REGION Network 15: Position Carrier Control First Carrier in Accumulation Zone
   RUNG wire#powerrail
      Contact( "EMS".Zone[#Zone].AccumZone )
      wire#w1
      I_Contact( "EMS".Zone[#NextZone].ZoneFull )
      wire#w2
      Move(in := #NextStopPosition, out1 => #TrafficCopCarrierZnBuffer[#ZonePos].CommandPos)
      wire#w3
      I_Contact( "EMS".Zone[#Zone].FinePosStopZone )
      Sub(in1 := #TrafficCopCarrierZnBuffer[#ZonePos].CommandPos, in2 := "EMS".CoarsePositionTolerance, out => #TrafficCopCarrierZnBuffer[#ZonePos].CommandPosLowLimit)
      Add(in1 := #TrafficCopCarrierZnBuffer[#ZonePos].CommandPos, in2 := "EMS".CoarsePositionTolerance, out => #TrafficCopCarrierZnBuffer[#ZonePos].CommandPosHighLimit)
   END_RUNG
   RUNG wire#w1
      { S7_Templates := "SrcType := DInt" } LT_Contact(in1 := "EMS".Zone[#Zone].CarrierZnStatus[#ZonePos].Position, in2 := #EndPos_LowLimit)
   END_RUNG wire#w2
   RUNG wire#w1
      { S7_Templates := "SrcType := DInt" } GE_Contact(in1 := "EMS".Zone[#Zone].CarrierZnStatus[#ZonePos].Position, in2 := #EndPos_LowLimit)
      { S7_Templates := "SrcType := DInt" } LE_Contact(in1 := "EMS".Zone[#Zone].CarrierZnStatus[#ZonePos].Position, in2 := #EndPos_HighLimit)
      { S7_Templates := "SrcType := Word" } EQ_Contact(in1 := "EMS".Zone[#NextZone].CarrierZnStatus[1].CarrierNumber, in2 := 0)
   END_RUNG wire#w2
   RUNG wire#powerrail
      Contact( "EMS".Zone[#Zone].ProductionZone )
      { S7_Templates := "SrcType := DInt" } LT_Contact(in1 := "EMS".Zone[#Zone].CarrierZnStatus[#ZonePos].Position, in2 := #ClrOfStopPos_LowLimit)
      Move(in := #ClearOfStopPos, out1 => #TrafficCopCarrierZnBuffer[#ZonePos].CommandPos)
   END_RUNG wire#w3
   RUNG wire#w3
      Contact( "EMS".Zone[#Zone].FinePosStopZone )
      Sub(in1 := #TrafficCopCarrierZnBuffer[#ZonePos].CommandPos, in2 := "EMS".FinePositionTolerance, out => #TrafficCopCarrierZnBuffer[#ZonePos].CommandPosLowLimit)
      Add(in1 := #TrafficCopCarrierZnBuffer[#ZonePos].CommandPos, in2 := "EMS".FinePositionTolerance, out => #TrafficCopCarrierZnBuffer[#ZonePos].CommandPosHighLimit)
   END_RUNG
   // the same network as SCL:
   #_w1 := "EMS".Zone[#Zone].AccumZone AND (NOT "EMS".Zone[#NextZone].ZoneFull OR ("EMS".Zone[#Zone].CarrierZnStatus[#ZonePos].Position < #EndPos_LowLimit) OR (("EMS".Zone[#Zone].CarrierZnStatus[#ZonePos].Position >= #EndPos_LowLimit) AND ("EMS".Zone[#Zone].CarrierZnStatus[#ZonePos].Position <= #EndPos_HighLimit) AND ("EMS".Zone[#NextZone].CarrierZnStatus[1].CarrierNumber = 0)));
   IF #_w1 THEN #TrafficCopCarrierZnBuffer[#ZonePos].CommandPos := #NextStopPosition; END_IF;
   #_w2 := "EMS".Zone[#Zone].ProductionZone AND ("EMS".Zone[#Zone].CarrierZnStatus[#ZonePos].Position < #ClrOfStopPos_LowLimit);
   IF #_w2 THEN #TrafficCopCarrierZnBuffer[#ZonePos].CommandPos := #ClearOfStopPos; END_IF;
   #_w3 := #_w1 OR #_w2;
   IF #_w3 AND NOT "EMS".Zone[#Zone].FinePosStopZone THEN
       #TrafficCopCarrierZnBuffer[#ZonePos].CommandPosLowLimit := #TrafficCopCarrierZnBuffer[#ZonePos].CommandPos - "EMS".CoarsePositionTolerance;
       #TrafficCopCarrierZnBuffer[#ZonePos].CommandPosHighLimit := #TrafficCopCarrierZnBuffer[#ZonePos].CommandPos + "EMS".CoarsePositionTolerance;
   END_IF;
   IF #_w3 AND "EMS".Zone[#Zone].FinePosStopZone THEN
       #TrafficCopCarrierZnBuffer[#ZonePos].CommandPosLowLimit := #TrafficCopCarrierZnBuffer[#ZonePos].CommandPos - "EMS".FinePositionTolerance;
       #TrafficCopCarrierZnBuffer[#ZonePos].CommandPosHighLimit := #TrafficCopCarrierZnBuffer[#ZonePos].CommandPos + "EMS".FinePositionTolerance;
   END_IF;
END_REGION

REGION Network 16: Position Carrier Control First Carrier in Production Zone
   // Control of First Carrier in Zone Closest to end position/Stop.  Move command is issued to carrier. Carrier will move in auto.
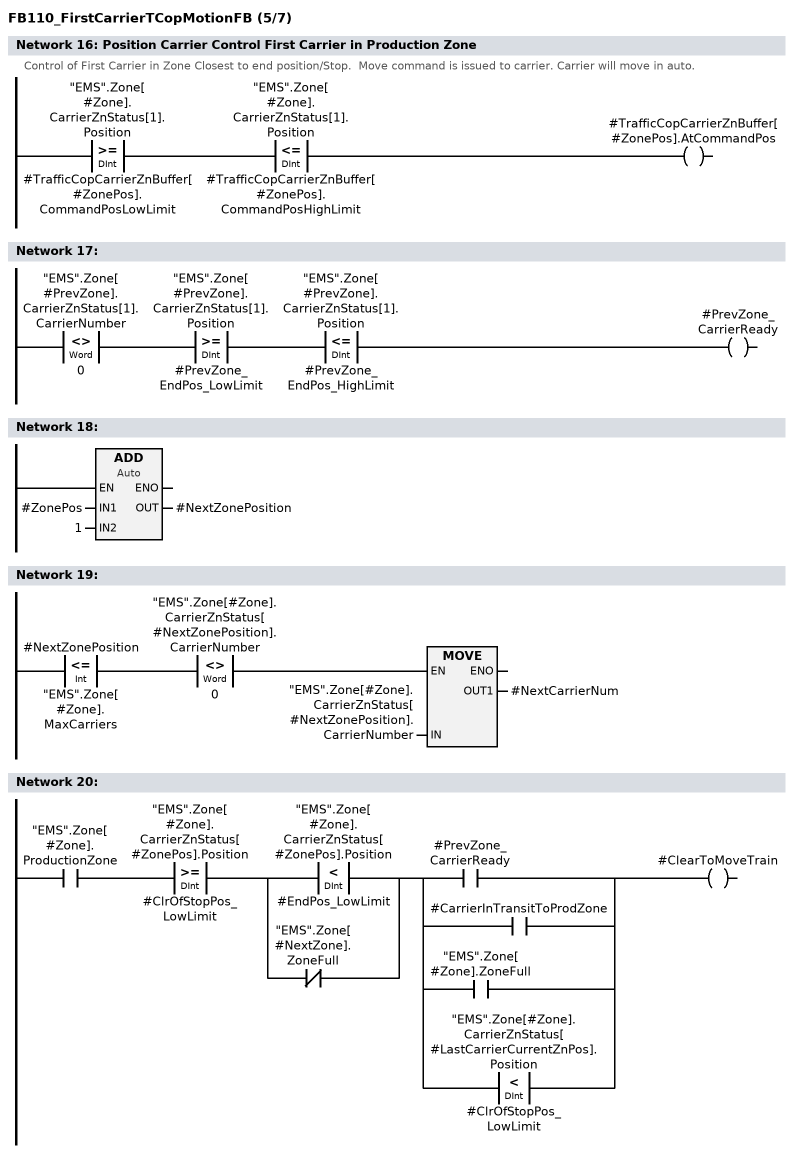
   RUNG wire#powerrail
      { S7_Templates := "SrcType := DInt" } GE_Contact(in1 := "EMS".Zone[#Zone].CarrierZnStatus[1].Position, in2 := #TrafficCopCarrierZnBuffer[#ZonePos].CommandPosLowLimit)
      { S7_Templates := "SrcType := DInt" } LE_Contact(in1 := "EMS".Zone[#Zone].CarrierZnStatus[1].Position, in2 := #TrafficCopCarrierZnBuffer[#ZonePos].CommandPosHighLimit)
      Coil( #TrafficCopCarrierZnBuffer[#ZonePos].AtCommandPos )
   END_RUNG
   // the same network as SCL:
   #TrafficCopCarrierZnBuffer[#ZonePos].AtCommandPos := ("EMS".Zone[#Zone].CarrierZnStatus[1].Position >= #TrafficCopCarrierZnBuffer[#ZonePos].CommandPosLowLimit) AND ("EMS".Zone[#Zone].CarrierZnStatus[1].Position <= #TrafficCopCarrierZnBuffer[#ZonePos].CommandPosHighLimit);
END_REGION

REGION Network 17
   RUNG wire#powerrail
      { S7_Templates := "SrcType := Word" } NE_Contact(in1 := "EMS".Zone[#PrevZone].CarrierZnStatus[1].CarrierNumber, in2 := 0)
      { S7_Templates := "SrcType := DInt" } GE_Contact(in1 := "EMS".Zone[#PrevZone].CarrierZnStatus[1].Position, in2 := #PrevZone_EndPos_LowLimit)
      { S7_Templates := "SrcType := DInt" } LE_Contact(in1 := "EMS".Zone[#PrevZone].CarrierZnStatus[1].Position, in2 := #PrevZone_EndPos_HighLimit)
      Coil( #PrevZone_CarrierReady )
   END_RUNG
   // the same network as SCL:
   #PrevZone_CarrierReady := ("EMS".Zone[#PrevZone].CarrierZnStatus[1].CarrierNumber <> 0) AND ("EMS".Zone[#PrevZone].CarrierZnStatus[1].Position >= #PrevZone_EndPos_LowLimit) AND ("EMS".Zone[#PrevZone].CarrierZnStatus[1].Position <= #PrevZone_EndPos_HighLimit);
END_REGION

REGION Network 18
   RUNG wire#powerrail
      Add(in1 := #ZonePos, in2 := 1, out => #NextZonePosition)
   END_RUNG
   // the same network as SCL:
   #NextZonePosition := #ZonePos + 1;
END_REGION

REGION Network 19
   RUNG wire#powerrail
      { S7_Templates := "SrcType := Int" } LE_Contact(in1 := #NextZonePosition, in2 := "EMS".Zone[#Zone].MaxCarriers)
      { S7_Templates := "SrcType := Word" } NE_Contact(in1 := "EMS".Zone[#Zone].CarrierZnStatus[#NextZonePosition].CarrierNumber, in2 := 0)
      Move(in := "EMS".Zone[#Zone].CarrierZnStatus[#NextZonePosition].CarrierNumber, out1 => #NextCarrierNum)
   END_RUNG
   // the same network as SCL:
   IF (#NextZonePosition <= "EMS".Zone[#Zone].MaxCarriers) AND ("EMS".Zone[#Zone].CarrierZnStatus[#NextZonePosition].CarrierNumber <> 0) THEN
       #NextCarrierNum := "EMS".Zone[#Zone].CarrierZnStatus[#NextZonePosition].CarrierNumber;
   END_IF;
END_REGION

REGION Network 20
   RUNG wire#powerrail
      Contact( "EMS".Zone[#Zone].ProductionZone )
      { S7_Templates := "SrcType := DInt" } GE_Contact(in1 := "EMS".Zone[#Zone].CarrierZnStatus[#ZonePos].Position, in2 := #ClrOfStopPos_LowLimit)
      wire#w1
      { S7_Templates := "SrcType := DInt" } LT_Contact(in1 := "EMS".Zone[#Zone].CarrierZnStatus[#ZonePos].Position, in2 := #EndPos_LowLimit)
      wire#w2
      Contact( #PrevZone_CarrierReady )
      wire#w3
      Coil( #ClearToMoveTrain )
   END_RUNG
   RUNG wire#w1
      I_Contact( "EMS".Zone[#NextZone].ZoneFull )
   END_RUNG wire#w2
   RUNG wire#w2
      Contact( #CarrierInTransitToProdZone )
   END_RUNG wire#w3
   RUNG wire#w2
      Contact( "EMS".Zone[#Zone].ZoneFull )
   END_RUNG wire#w3
   RUNG wire#w2
      { S7_Templates := "SrcType := DInt" } LT_Contact(in1 := "EMS".Zone[#Zone].CarrierZnStatus[#LastCarrierCurrentZnPos].Position, in2 := #ClrOfStopPos_LowLimit)
   END_RUNG wire#w3
   // the same network as SCL:
   #ClearToMoveTrain := "EMS".Zone[#Zone].ProductionZone AND ("EMS".Zone[#Zone].CarrierZnStatus[#ZonePos].Position >= #ClrOfStopPos_LowLimit) AND (("EMS".Zone[#Zone].CarrierZnStatus[#ZonePos].Position < #EndPos_LowLimit) OR NOT "EMS".Zone[#NextZone].ZoneFull) AND (#PrevZone_CarrierReady OR #CarrierInTransitToProdZone OR "EMS".Zone[#Zone].ZoneFull OR ("EMS".Zone[#Zone].CarrierZnStatus[#LastCarrierCurrentZnPos].Position < #ClrOfStopPos_LowLimit));
END_REGION

REGION Network 21
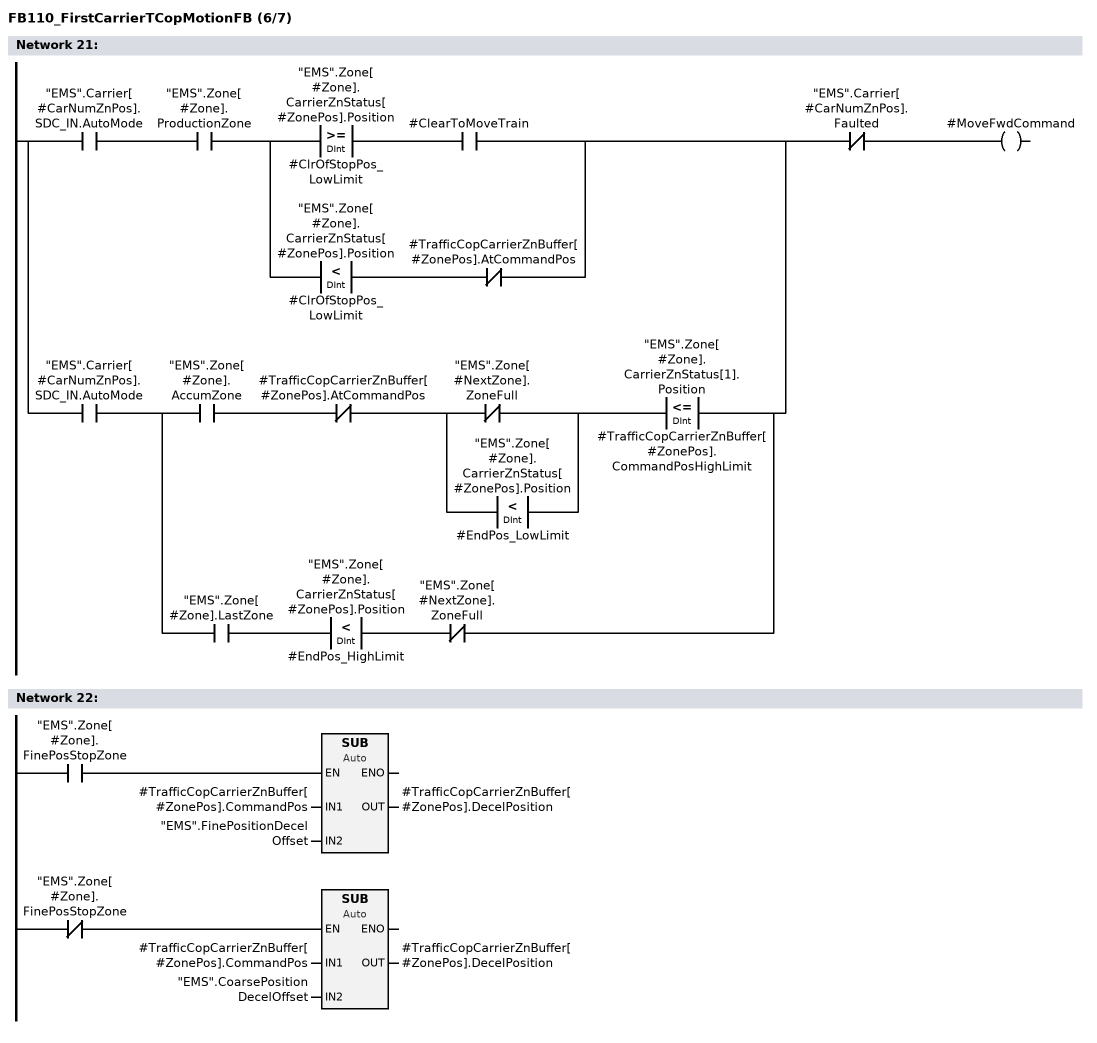
   RUNG wire#powerrail
      Contact( "EMS".Carrier[#CarNumZnPos].SDC_IN.AutoMode )
      Contact( "EMS".Zone[#Zone].ProductionZone )
      wire#w1
      { S7_Templates := "SrcType := DInt" } GE_Contact(in1 := "EMS".Zone[#Zone].CarrierZnStatus[#ZonePos].Position, in2 := #ClrOfStopPos_LowLimit)
      Contact( #ClearToMoveTrain )
      wire#w2
      I_Contact( "EMS".Carrier[#CarNumZnPos].Faulted )
      Coil( #MoveFwdCommand )
   END_RUNG
   RUNG wire#w1
      { S7_Templates := "SrcType := DInt" } LT_Contact(in1 := "EMS".Zone[#Zone].CarrierZnStatus[#ZonePos].Position, in2 := #ClrOfStopPos_LowLimit)
      I_Contact( #TrafficCopCarrierZnBuffer[#ZonePos].AtCommandPos )
   END_RUNG wire#w2
   RUNG wire#powerrail
      Contact( "EMS".Carrier[#CarNumZnPos].SDC_IN.AutoMode )
      wire#w3
      Contact( "EMS".Zone[#Zone].AccumZone )
      I_Contact( #TrafficCopCarrierZnBuffer[#ZonePos].AtCommandPos )
      wire#w4
      I_Contact( "EMS".Zone[#NextZone].ZoneFull )
      wire#w5
      { S7_Templates := "SrcType := DInt" } LE_Contact(in1 := "EMS".Zone[#Zone].CarrierZnStatus[1].Position, in2 := #TrafficCopCarrierZnBuffer[#ZonePos].CommandPosHighLimit)
   END_RUNG wire#w2
   RUNG wire#w4
      { S7_Templates := "SrcType := DInt" } LT_Contact(in1 := "EMS".Zone[#Zone].CarrierZnStatus[#ZonePos].Position, in2 := #EndPos_LowLimit)
   END_RUNG wire#w5
   RUNG wire#w3
      Contact( "EMS".Zone[#Zone].LastZone )
      { S7_Templates := "SrcType := DInt" } LT_Contact(in1 := "EMS".Zone[#Zone].CarrierZnStatus[#ZonePos].Position, in2 := #EndPos_HighLimit)
      I_Contact( "EMS".Zone[#NextZone].ZoneFull )
   END_RUNG wire#w2
   // the same network as SCL:
   #MoveFwdCommand := (("EMS".Carrier[#CarNumZnPos].SDC_IN.AutoMode AND "EMS".Zone[#Zone].ProductionZone AND ((("EMS".Zone[#Zone].CarrierZnStatus[#ZonePos].Position >= #ClrOfStopPos_LowLimit) AND #ClearToMoveTrain) OR (("EMS".Zone[#Zone].CarrierZnStatus[#ZonePos].Position < #ClrOfStopPos_LowLimit) AND NOT #TrafficCopCarrierZnBuffer[#ZonePos].AtCommandPos))) OR ("EMS".Carrier[#CarNumZnPos].SDC_IN.AutoMode AND (("EMS".Zone[#Zone].AccumZone AND NOT #TrafficCopCarrierZnBuffer[#ZonePos].AtCommandPos AND (NOT "EMS".Zone[#NextZone].ZoneFull OR ("EMS".Zone[#Zone].CarrierZnStatus[#ZonePos].Position < #EndPos_LowLimit)) AND ("EMS".Zone[#Zone].CarrierZnStatus[1].Position <= #TrafficCopCarrierZnBuffer[#ZonePos].CommandPosHighLimit)) OR ("EMS".Zone[#Zone].LastZone AND ("EMS".Zone[#Zone].CarrierZnStatus[#ZonePos].Position < #EndPos_HighLimit) AND NOT "EMS".Zone[#NextZone].ZoneFull)))) AND NOT "EMS".Carrier[#CarNumZnPos].Faulted;
END_REGION

REGION Network 22
   RUNG wire#powerrail
      Contact( "EMS".Zone[#Zone].FinePosStopZone )
      Sub(in1 := #TrafficCopCarrierZnBuffer[#ZonePos].CommandPos, in2 := "EMS".FinePositionDecelOffset, out => #TrafficCopCarrierZnBuffer[#ZonePos].DecelPosition)
   END_RUNG
   RUNG wire#powerrail
      I_Contact( "EMS".Zone[#Zone].FinePosStopZone )
      Sub(in1 := #TrafficCopCarrierZnBuffer[#ZonePos].CommandPos, in2 := "EMS".CoarsePositionDecelOffset, out => #TrafficCopCarrierZnBuffer[#ZonePos].DecelPosition)
   END_RUNG
   // the same network as SCL:
   IF "EMS".Zone[#Zone].FinePosStopZone THEN
       #TrafficCopCarrierZnBuffer[#ZonePos].DecelPosition := #TrafficCopCarrierZnBuffer[#ZonePos].CommandPos - "EMS".FinePositionDecelOffset;
   END_IF;
   IF NOT "EMS".Zone[#Zone].FinePosStopZone THEN
       #TrafficCopCarrierZnBuffer[#ZonePos].DecelPosition := #TrafficCopCarrierZnBuffer[#ZonePos].CommandPos - "EMS".CoarsePositionDecelOffset;
   END_IF;
END_REGION

REGION Network 23
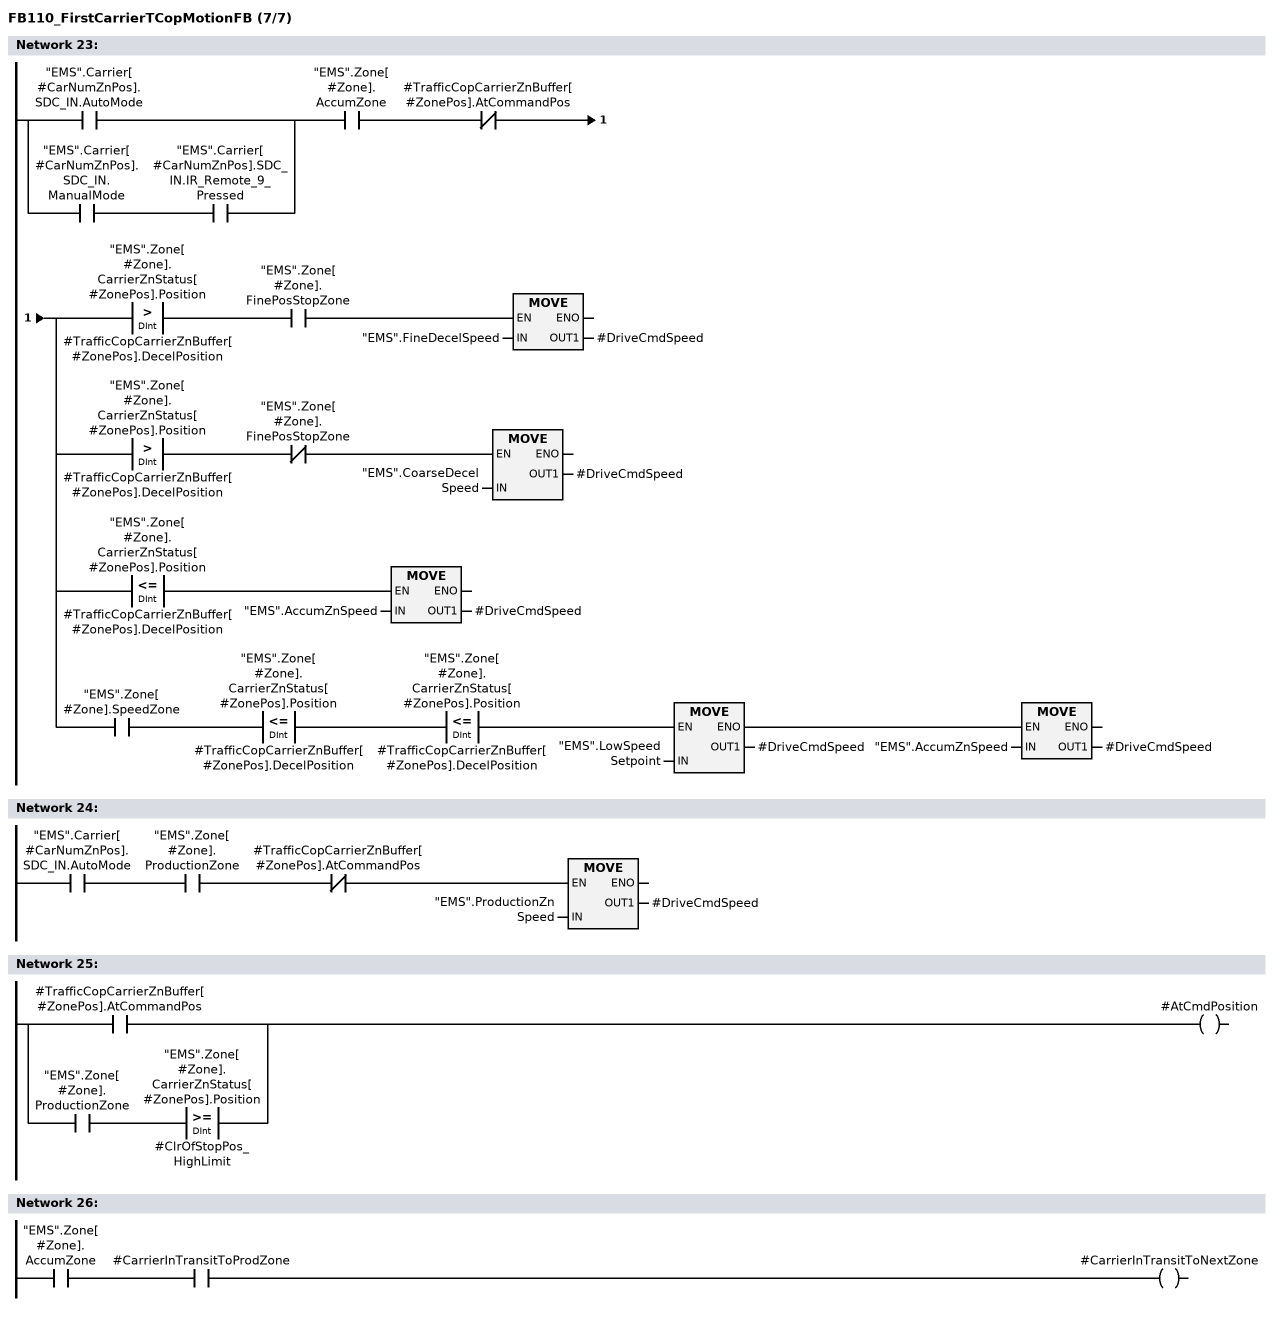
   RUNG wire#powerrail
      Contact( "EMS".Carrier[#CarNumZnPos].SDC_IN.AutoMode )
      wire#w1
      Contact( "EMS".Zone[#Zone].AccumZone )
      I_Contact( #TrafficCopCarrierZnBuffer[#ZonePos].AtCommandPos )
      wire#w2
      { S7_Templates := "SrcType := DInt" } GT_Contact(in1 := "EMS".Zone[#Zone].CarrierZnStatus[#ZonePos].Position, in2 := #TrafficCopCarrierZnBuffer[#ZonePos].DecelPosition)
      Contact( "EMS".Zone[#Zone].FinePosStopZone )
      Move(in := "EMS".FineDecelSpeed, out1 => #DriveCmdSpeed)
   END_RUNG
   RUNG wire#powerrail
      Contact( "EMS".Carrier[#CarNumZnPos].SDC_IN.ManualMode )
      Contact( "EMS".Carrier[#CarNumZnPos].SDC_IN.IR_Remote_9_Pressed )
   END_RUNG wire#w1
   RUNG wire#w2
      { S7_Templates := "SrcType := DInt" } GT_Contact(in1 := "EMS".Zone[#Zone].CarrierZnStatus[#ZonePos].Position, in2 := #TrafficCopCarrierZnBuffer[#ZonePos].DecelPosition)
      I_Contact( "EMS".Zone[#Zone].FinePosStopZone )
      Move(in := "EMS".CoarseDecelSpeed, out1 => #DriveCmdSpeed)
   END_RUNG
   RUNG wire#w2
      { S7_Templates := "SrcType := DInt" } LE_Contact(in1 := "EMS".Zone[#Zone].CarrierZnStatus[#ZonePos].Position, in2 := #TrafficCopCarrierZnBuffer[#ZonePos].DecelPosition)
      Move(in := "EMS".AccumZnSpeed, out1 => #DriveCmdSpeed)
   END_RUNG
   RUNG wire#w2
      Contact( "EMS".Zone[#Zone].SpeedZone )
      { S7_Templates := "SrcType := DInt" } LE_Contact(in1 := "EMS".Zone[#Zone].CarrierZnStatus[#ZonePos].Position, in2 := #TrafficCopCarrierZnBuffer[#ZonePos].DecelPosition)
      { S7_Templates := "SrcType := DInt" } LE_Contact(in1 := "EMS".Zone[#Zone].CarrierZnStatus[#ZonePos].Position, in2 := #TrafficCopCarrierZnBuffer[#ZonePos].DecelPosition)
      Move(in := "EMS".LowSpeedSetpoint, out1 => #DriveCmdSpeed)
      Move(in := "EMS".AccumZnSpeed, out1 => #DriveCmdSpeed)
   END_RUNG
   // the same network as SCL:
   #_w1 := ("EMS".Carrier[#CarNumZnPos].SDC_IN.AutoMode OR ("EMS".Carrier[#CarNumZnPos].SDC_IN.ManualMode AND "EMS".Carrier[#CarNumZnPos].SDC_IN.IR_Remote_9_Pressed)) AND "EMS".Zone[#Zone].AccumZone AND NOT #TrafficCopCarrierZnBuffer[#ZonePos].AtCommandPos;
   IF #_w1 AND ("EMS".Zone[#Zone].CarrierZnStatus[#ZonePos].Position > #TrafficCopCarrierZnBuffer[#ZonePos].DecelPosition) AND "EMS".Zone[#Zone].FinePosStopZone THEN
       #DriveCmdSpeed := "EMS".FineDecelSpeed;
   END_IF;
   IF #_w1 AND ("EMS".Zone[#Zone].CarrierZnStatus[#ZonePos].Position > #TrafficCopCarrierZnBuffer[#ZonePos].DecelPosition) AND NOT "EMS".Zone[#Zone].FinePosStopZone THEN
       #DriveCmdSpeed := "EMS".CoarseDecelSpeed;
   END_IF;
   IF #_w1 AND ("EMS".Zone[#Zone].CarrierZnStatus[#ZonePos].Position <= #TrafficCopCarrierZnBuffer[#ZonePos].DecelPosition) THEN
       #DriveCmdSpeed := "EMS".AccumZnSpeed;
   END_IF;
   IF #_w1 AND "EMS".Zone[#Zone].SpeedZone AND ("EMS".Zone[#Zone].CarrierZnStatus[#ZonePos].Position <= #TrafficCopCarrierZnBuffer[#ZonePos].DecelPosition) AND ("EMS".Zone[#Zone].CarrierZnStatus[#ZonePos].Position <= #TrafficCopCarrierZnBuffer[#ZonePos].DecelPosition) THEN
       #DriveCmdSpeed := "EMS".LowSpeedSetpoint;
       #DriveCmdSpeed := "EMS".AccumZnSpeed;
   END_IF;
END_REGION

REGION Network 24
   RUNG wire#powerrail
      Contact( "EMS".Carrier[#CarNumZnPos].SDC_IN.AutoMode )
      Contact( "EMS".Zone[#Zone].ProductionZone )
      I_Contact( #TrafficCopCarrierZnBuffer[#ZonePos].AtCommandPos )
      Move(in := "EMS".ProductionZnSpeed, out1 => #DriveCmdSpeed)
   END_RUNG
   // the same network as SCL:
   IF "EMS".Carrier[#CarNumZnPos].SDC_IN.AutoMode AND "EMS".Zone[#Zone].ProductionZone AND NOT #TrafficCopCarrierZnBuffer[#ZonePos].AtCommandPos THEN
       #DriveCmdSpeed := "EMS".ProductionZnSpeed;
   END_IF;
END_REGION

REGION Network 25
   RUNG wire#powerrail
      Contact( #TrafficCopCarrierZnBuffer[#ZonePos].AtCommandPos )
      wire#w1
      Coil( #AtCmdPosition )
   END_RUNG
   RUNG wire#powerrail
      Contact( "EMS".Zone[#Zone].ProductionZone )
      { S7_Templates := "SrcType := DInt" } GE_Contact(in1 := "EMS".Zone[#Zone].CarrierZnStatus[#ZonePos].Position, in2 := #ClrOfStopPos_HighLimit)
   END_RUNG wire#w1
   // the same network as SCL:
   #AtCmdPosition := #TrafficCopCarrierZnBuffer[#ZonePos].AtCommandPos OR ("EMS".Zone[#Zone].ProductionZone AND ("EMS".Zone[#Zone].CarrierZnStatus[#ZonePos].Position >= #ClrOfStopPos_HighLimit));
END_REGION

REGION Network 26
   RUNG wire#powerrail
      Contact( "EMS".Zone[#Zone].AccumZone )
      Contact( #CarrierInTransitToProdZone )
      Coil( #CarrierInTransitToNextZone )
   END_RUNG
   // the same network as SCL:
   #CarrierInTransitToNextZone := "EMS".Zone[#Zone].AccumZone AND #CarrierInTransitToProdZone;
END_REGION
END_FUNCTION_BLOCK

FUNCTION_BLOCK "FB111_NextCarrierTCopMotionFB"   // FB111, LAD
{ S7_Optimized_Access := 'TRUE' }
VERSION : 0.1
   VAR_INPUT
      Zone : Int;
      ZonePos : Int;
   END_VAR
   VAR_OUTPUT
      CarrierNumber : Int;
      MoveFwdCommand : Bool;
      DriveCmdSpeed : Int;
      NextStopPosition : DWord;
      NextCarrierNum : Word;
      AtCmdPosition : Bool;
   END_VAR
   VAR
      LowSpeedSetpoint : Word;
      HighSpeedSetpoint : Word;
      TrafficCopCarrierZnBuffer : Array[0..40] of "UDT_TrafficCop";
      NextZonePosition : Int;
      PreviousZoneCarNum : Int;
      PrevZonePos : Int;
      CarrNumNextZn : Int;
      PreviousCarrPos : DWord;
      CarNumZnPos : Int;
   END_VAR
   VAR_TEMP   // added for the SCL form of the ladder/FBD networks
      _w1 : Bool;
   END_VAR
BEGIN

REGION Network 1
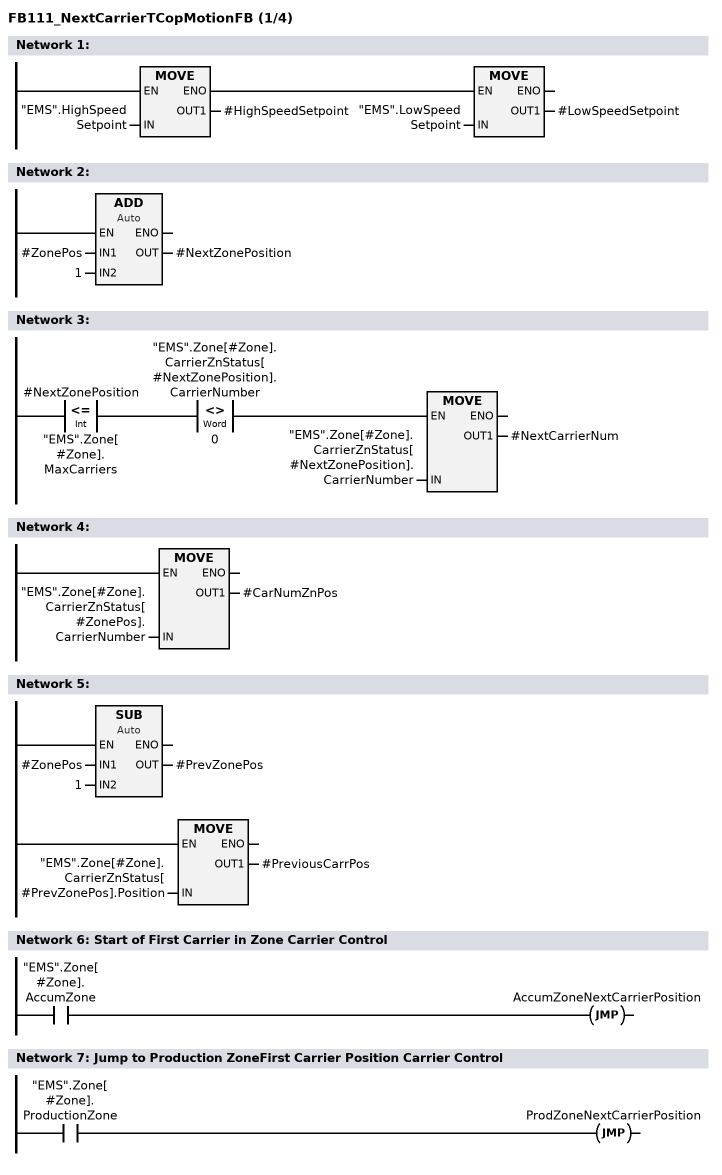
   RUNG wire#powerrail
      Move(in := "EMS".HighSpeedSetpoint, out1 => #HighSpeedSetpoint)
      Move(in := "EMS".LowSpeedSetpoint, out1 => #LowSpeedSetpoint)
   END_RUNG
   // the same network as SCL:
   #HighSpeedSetpoint := "EMS".HighSpeedSetpoint;
   #LowSpeedSetpoint := "EMS".LowSpeedSetpoint;
END_REGION

REGION Network 2
   RUNG wire#powerrail
      Add(in1 := #ZonePos, in2 := 1, out => #NextZonePosition)
   END_RUNG
   // the same network as SCL:
   #NextZonePosition := #ZonePos + 1;
END_REGION

REGION Network 3
   RUNG wire#powerrail
      { S7_Templates := "SrcType := Int" } LE_Contact(in1 := #NextZonePosition, in2 := "EMS".Zone[#Zone].MaxCarriers)
      { S7_Templates := "SrcType := Word" } NE_Contact(in1 := "EMS".Zone[#Zone].CarrierZnStatus[#NextZonePosition].CarrierNumber, in2 := 0)
      Move(in := "EMS".Zone[#Zone].CarrierZnStatus[#NextZonePosition].CarrierNumber, out1 => #NextCarrierNum)
   END_RUNG
   // the same network as SCL:
   IF (#NextZonePosition <= "EMS".Zone[#Zone].MaxCarriers) AND ("EMS".Zone[#Zone].CarrierZnStatus[#NextZonePosition].CarrierNumber <> 0) THEN
       #NextCarrierNum := "EMS".Zone[#Zone].CarrierZnStatus[#NextZonePosition].CarrierNumber;
   END_IF;
END_REGION

REGION Network 4
   RUNG wire#powerrail
      Move(in := "EMS".Zone[#Zone].CarrierZnStatus[#ZonePos].CarrierNumber, out1 => #CarNumZnPos)
   END_RUNG
   // the same network as SCL:
   #CarNumZnPos := "EMS".Zone[#Zone].CarrierZnStatus[#ZonePos].CarrierNumber;
END_REGION

REGION Network 5
   RUNG wire#powerrail
      Sub(in1 := #ZonePos, in2 := 1, out => #PrevZonePos)
   END_RUNG
   RUNG wire#powerrail
      Move(in := "EMS".Zone[#Zone].CarrierZnStatus[#PrevZonePos].Position, out1 => #PreviousCarrPos)
   END_RUNG
   // the same network as SCL:
   #PrevZonePos := #ZonePos - 1;
   #PreviousCarrPos := "EMS".Zone[#Zone].CarrierZnStatus[#PrevZonePos].Position;
END_REGION

REGION Network 6: Start of First Carrier in Zone Carrier Control
   RUNG wire#powerrail
      Contact( "EMS".Zone[#Zone].AccumZone )
      JumpCoil( AccumZoneNextCarrierPosition )
   END_RUNG
   // the same network as SCL:
   IF "EMS".Zone[#Zone].AccumZone THEN GOTO AccumZoneNextCarrierPosition; END_IF;
END_REGION

REGION Network 7: Jump to Production ZoneFirst Carrier Position Carrier Control
   RUNG wire#powerrail
      Contact( "EMS".Zone[#Zone].ProductionZone )
      JumpCoil( ProdZoneNextCarrierPosition )
   END_RUNG
   // the same network as SCL:
   IF "EMS".Zone[#Zone].ProductionZone THEN GOTO ProdZoneNextCarrierPosition; END_IF;
END_REGION

REGION Network 8: Position Carrier Control First Carrier in Accumulation Zone
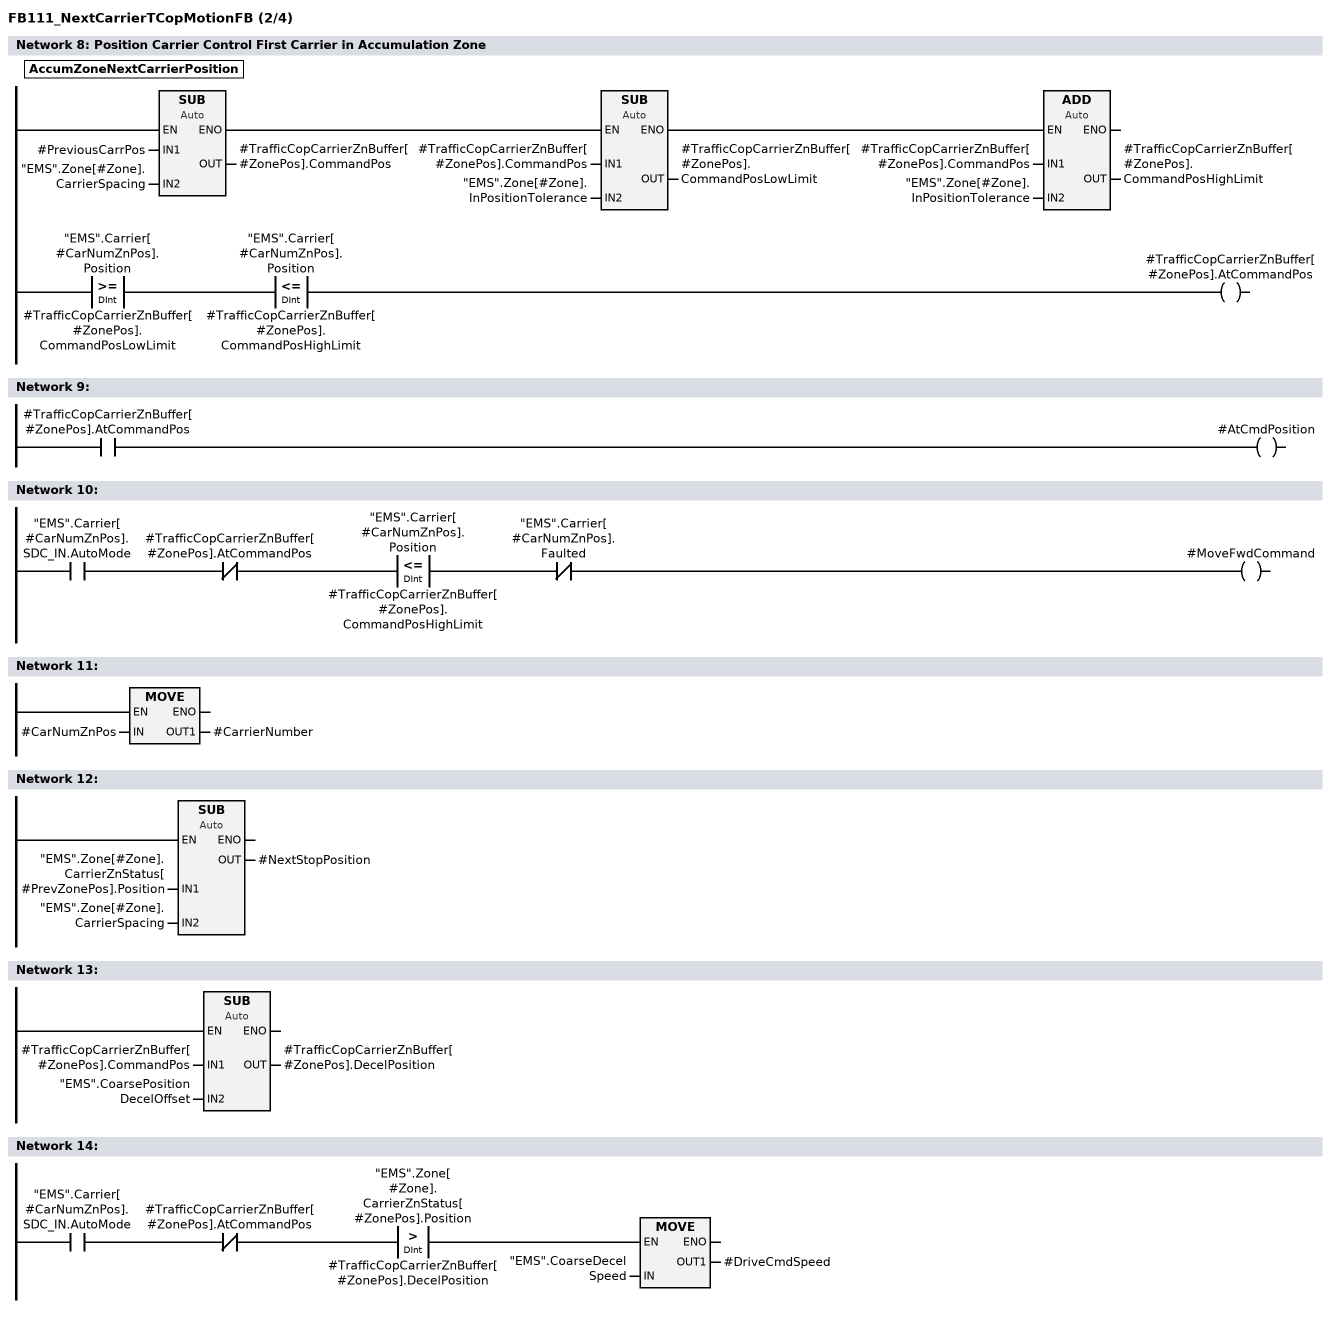
   Label( AccumZoneNextCarrierPosition )
   RUNG wire#powerrail
      Sub(in1 := #PreviousCarrPos, in2 := "EMS".Zone[#Zone].CarrierSpacing, out => #TrafficCopCarrierZnBuffer[#ZonePos].CommandPos)
      Sub(in1 := #TrafficCopCarrierZnBuffer[#ZonePos].CommandPos, in2 := "EMS".Zone[#Zone].InPositionTolerance, out => #TrafficCopCarrierZnBuffer[#ZonePos].CommandPosLowLimit)
      Add(in1 := #TrafficCopCarrierZnBuffer[#ZonePos].CommandPos, in2 := "EMS".Zone[#Zone].InPositionTolerance, out => #TrafficCopCarrierZnBuffer[#ZonePos].CommandPosHighLimit)
   END_RUNG
   RUNG wire#powerrail
      { S7_Templates := "SrcType := DInt" } GE_Contact(in1 := "EMS".Carrier[#CarNumZnPos].Position, in2 := #TrafficCopCarrierZnBuffer[#ZonePos].CommandPosLowLimit)
      { S7_Templates := "SrcType := DInt" } LE_Contact(in1 := "EMS".Carrier[#CarNumZnPos].Position, in2 := #TrafficCopCarrierZnBuffer[#ZonePos].CommandPosHighLimit)
      Coil( #TrafficCopCarrierZnBuffer[#ZonePos].AtCommandPos )
   END_RUNG
   // the same network as SCL:
   AccumZoneNextCarrierPosition:
   #TrafficCopCarrierZnBuffer[#ZonePos].CommandPos := #PreviousCarrPos - "EMS".Zone[#Zone].CarrierSpacing;
   #TrafficCopCarrierZnBuffer[#ZonePos].CommandPosLowLimit := #TrafficCopCarrierZnBuffer[#ZonePos].CommandPos - "EMS".Zone[#Zone].InPositionTolerance;
   #TrafficCopCarrierZnBuffer[#ZonePos].CommandPosHighLimit := #TrafficCopCarrierZnBuffer[#ZonePos].CommandPos + "EMS".Zone[#Zone].InPositionTolerance;
   #TrafficCopCarrierZnBuffer[#ZonePos].AtCommandPos := ("EMS".Carrier[#CarNumZnPos].Position >= #TrafficCopCarrierZnBuffer[#ZonePos].CommandPosLowLimit) AND ("EMS".Carrier[#CarNumZnPos].Position <= #TrafficCopCarrierZnBuffer[#ZonePos].CommandPosHighLimit);
END_REGION

REGION Network 9
   RUNG wire#powerrail
      Contact( #TrafficCopCarrierZnBuffer[#ZonePos].AtCommandPos )
      Coil( #AtCmdPosition )
   END_RUNG
   // the same network as SCL:
   #AtCmdPosition := #TrafficCopCarrierZnBuffer[#ZonePos].AtCommandPos;
END_REGION

REGION Network 10
   RUNG wire#powerrail
      Contact( "EMS".Carrier[#CarNumZnPos].SDC_IN.AutoMode )
      I_Contact( #TrafficCopCarrierZnBuffer[#ZonePos].AtCommandPos )
      { S7_Templates := "SrcType := DInt" } LE_Contact(in1 := "EMS".Carrier[#CarNumZnPos].Position, in2 := #TrafficCopCarrierZnBuffer[#ZonePos].CommandPosHighLimit)
      I_Contact( "EMS".Carrier[#CarNumZnPos].Faulted )
      Coil( #MoveFwdCommand )
   END_RUNG
   // the same network as SCL:
   #MoveFwdCommand := "EMS".Carrier[#CarNumZnPos].SDC_IN.AutoMode AND NOT #TrafficCopCarrierZnBuffer[#ZonePos].AtCommandPos AND ("EMS".Carrier[#CarNumZnPos].Position <= #TrafficCopCarrierZnBuffer[#ZonePos].CommandPosHighLimit) AND NOT "EMS".Carrier[#CarNumZnPos].Faulted;
END_REGION

REGION Network 11
   RUNG wire#powerrail
      Move(in := #CarNumZnPos, out1 => #CarrierNumber)
   END_RUNG
   // the same network as SCL:
   #CarrierNumber := #CarNumZnPos;
END_REGION
